   "TT426_4S_ALM_ANALOG_DB_LOW LEVEL VALUE (L)" : Real = PLC TT426_4S_ALM_ANALOG_DB."LOW LEVEL VALUE (L)" AT %DB2080.DBD26, 1 s
   "PIT424PORT_ALM_ANALOG_DB_HIGH LEVEL VALUE (H)" : Real = PLC PIT424PORT_ALM_ANALOG_DB."HIGH LEVEL VALUE (H)" AT %DB2070.DBD30, 1 s
   "TT426_4S_ALM_ANALOG_DB_VERY HIGH LEVEL VALUE (HH)" : Real = PLC TT426_4S_ALM_ANALOG_DB."VERY HIGH LEVEL VALUE (HH)" AT %DB2080.DBD34, 1 s
   "PT415_RIO7_ALM_ANALOG_DB_LOW LEVEL VALUE (L)" : Real = PLC PT415_RIO7_ALM_ANALOG_DB."LOW LEVEL VALUE (L)" AT %DB2225.DBD26, 1 s
   "PT415_RIO6_ALM_ANALOG_DB_VERY HIGH LEVEL VALUE (HH)" : Real = PLC PT415_RIO6_ALM_ANALOG_DB."VERY HIGH LEVEL VALUE (HH)" AT %DB2218.DBD34, 1 s
   "Sequence Times_DB_Pre-Dwell Timer_Days Left" : DInt = PLC "Sequence Times_DB"."Pre-Dwell Timer"."Days Left", 1 s
   "504_Tank Grouping_DB2020_Cycle Period_ET" : Time = PLC "504_Tank Grouping_DB2020"."Cycle Period".ET, 1 s
   "504_Tank Grouping_DB2020_Cycle Length_ET" : Time = PLC "504_Tank Grouping_DB2020"."Cycle Length".ET, 1 s
   "504_Tank Grouping_DB2020_Valve Cycle_Enable" : Bool = PLC "504_Tank Grouping_DB2020"."Valve Cycle".Enable, 1 s
   "504_Tank Grouping_DB2020_Valve Cycle_Period" : Time = PLC "504_Tank Grouping_DB2020"."Valve Cycle".Period, 1 s
   "504_Tank Grouping_DB2020_Valve Cycle_Length" : Time = PLC "504_Tank Grouping_DB2020"."Valve Cycle".Length, 1 s
   "Process Gas Compressor Running/Stopped" : Bool = PLC "Process Gas Compressor Running/Stopped" AT %I139.0, 1 s
   "PT415_FPT_ALM_ANALOG_DB_VERY LOW LEVEL VALUE (LL)" : Real = PLC PT415_FPT_ALM_ANALOG_DB."VERY LOW LEVEL VALUE (LL)" AT %DB2213.DBD22, 1 s
   "PT415_FPT_ALM_ANALOG_DB_LOW LEVEL VALUE (L)" : Real = PLC PT415_FPT_ALM_ANALOG_DB."LOW LEVEL VALUE (L)" AT %DB2213.DBD26, 1 s
   "PT415_FPT_ALM_ANALOG_DB_HIGH LEVEL VALUE (H)" : Real = PLC PT415_FPT_ALM_ANALOG_DB."HIGH LEVEL VALUE (H)" AT %DB2213.DBD30, 1 s
   "PT415_RIO7_ALM_ANALOG_DB_VERY LOW LEVEL VALUE (LL)" : Real = PLC PT415_RIO7_ALM_ANALOG_DB."VERY LOW LEVEL VALUE (LL)" AT %DB2225.DBD22, 1 s
   "PT415_FPT_ALM_ANALOG_DB_VERY HIGH LEVEL VALUE (HH)" : Real = PLC PT415_FPT_ALM_ANALOG_DB."VERY HIGH LEVEL VALUE (HH)" AT %DB2213.DBD34, 1 s
   "PT415_RIO3_ALM_ANALOG_DB_LOW LEVEL VALUE (L)" : Real = PLC PT415_RIO3_ALM_ANALOG_DB."LOW LEVEL VALUE (L)" AT %DB2215.DBD26, 1 s
   "PT415_RIO3_ALM_ANALOG_DB_HIGH LEVEL VALUE (H)" : Real = PLC PT415_RIO3_ALM_ANALOG_DB."HIGH LEVEL VALUE (H)" AT %DB2215.DBD30, 1 s
   "PT415_RIO3_ALM_ANALOG_DB_VERY HIGH LEVEL VALUE (HH)" : Real = PLC PT415_RIO3_ALM_ANALOG_DB."VERY HIGH LEVEL VALUE (HH)" AT %DB2215.DBD34, 1 s
   "PT415_RIO5_ALM_ANALOG_DB_VERY LOW LEVEL VALUE (LL)" : Real = PLC PT415_RIO5_ALM_ANALOG_DB."VERY LOW LEVEL VALUE (LL)" AT %DB2217.DBD22, 1 s
   "PT415_RIO5_ALM_ANALOG_DB_LOW LEVEL VALUE (L)" : Real = PLC PT415_RIO5_ALM_ANALOG_DB."LOW LEVEL VALUE (L)" AT %DB2217.DBD26, 1 s
   "PT415_RIO5_ALM_ANALOG_DB_HIGH LEVEL VALUE (H)" : Real = PLC PT415_RIO5_ALM_ANALOG_DB."HIGH LEVEL VALUE (H)" AT %DB2217.DBD30, 1 s
   "PT415_RIO5_ALM_ANALOG_DB_VERY HIGH LEVEL VALUE (HH)" : Real = PLC PT415_RIO5_ALM_ANALOG_DB."VERY HIGH LEVEL VALUE (HH)" AT %DB2217.DBD34, 1 s
   "PT415_RIO6_ALM_ANALOG_DB_VERY LOW LEVEL VALUE (LL)" : Real = PLC PT415_RIO6_ALM_ANALOG_DB."VERY LOW LEVEL VALUE (LL)" AT %DB2218.DBD22, 1 s
   "PT415_RIO6_ALM_ANALOG_DB_LOW LEVEL VALUE (L)" : Real = PLC PT415_RIO6_ALM_ANALOG_DB."LOW LEVEL VALUE (L)" AT %DB2218.DBD26, 1 s
   "PT415_RIO6_ALM_ANALOG_DB_HIGH LEVEL VALUE (H)" : Real = PLC PT415_RIO6_ALM_ANALOG_DB."HIGH LEVEL VALUE (H)" AT %DB2218.DBD30, 1 s
   "PT415_RIO3_ALM_ANALOG_DB_VERY LOW LEVEL VALUE (LL)" : Real = PLC PT415_RIO3_ALM_ANALOG_DB."VERY LOW LEVEL VALUE (LL)" AT %DB2215.DBD22, 1 s
   "RIO3_SPR_DI_33_4" : Bool = PLC RIO3_SPR_DI_33_4 AT %I33.4, 1 s
   "TT426_1S_ALM_ANALOG_DB_LOW LEVEL VALUE (L)" : Real = PLC TT426_1S_ALM_ANALOG_DB."LOW LEVEL VALUE (L)" AT %DB2076.DBD26, 1 s
   "TT426_1S_ALM_ANALOG_DB_VERY HIGH LEVEL VALUE (HH)" : Real = PLC TT426_1S_ALM_ANALOG_DB."VERY HIGH LEVEL VALUE (HH)" AT %DB2076.DBD34, 1 s
   "RIO6_SPR_DI_66_7" : Bool = PLC RIO6_SPR_DI_66_7 AT %I66.7, 1 s
   "RIO6_SPR_DI_66_5" : Bool = PLC RIO6_SPR_DI_66_5 AT %I66.5, 1 s
   "RIO6_SPR_DI_66_4" : Bool = PLC RIO6_SPR_DI_66_4 AT %I66.4, 1 s
   "RIO6_SPR_DI_66_3" : Bool = PLC RIO6_SPR_DI_66_3 AT %I66.3, 1 s
   "Tank 6S BWT Level High High Switch" : Bool = PLC "Tank 6S BWT Level High High Switch" AT %I66.2, 1 s
   "RIO6 Tanks Pressure Switch Hi Hi" : Bool = PLC "RIO6 Tanks Pressure Switch Hi Hi" AT %I66.1, 1 s
   "Tank 6P BWT Level High High Switch" : Bool = PLC "Tank 6P BWT Level High High Switch" AT %I66.0, 1 s
   "RIO6_SPR_DI_63_7" : Bool = PLC RIO6_SPR_DI_63_7 AT %I63.7, 1 s
   "RIO6_SPR_DI_63_6" : Bool = PLC RIO6_SPR_DI_63_6 AT %I63.6, 1 s
   "Tank 6S Tank Vent Valve 2 Feedback - Closed" : Bool = PLC "Tank 6S Tank Vent Valve 2 Feedback - Closed" AT %I63.5, 1 s
   "Tank 6S Tank Vent Valve 2 Feedback - Opened" : Bool = PLC "Tank 6S Tank Vent Valve 2 Feedback - Opened" AT %I63.4, 1 s
   "Tank 6S Tank Vent Valve 1 Feedback - Closed" : Bool = PLC "Tank 6S Tank Vent Valve 1 Feedback - Closed" AT %I63.3, 1 s
   "Tank 6S Tank Vent Valve 1 Feedback - Opened" : Bool = PLC "Tank 6S Tank Vent Valve 1 Feedback - Opened" AT %I63.2, 1 s
   "Tank 6S GTT Isolation Valve Feedback - Closed" : Bool = PLC "Tank 6S GTT Isolation Valve Feedback - Closed" AT %I63.1, 1 s
   "Tank 6S GTT Isolation Valve Feedback - Opened" : Bool = PLC "Tank 6S GTT Isolation Valve Feedback - Opened" AT %I63.0, 1 s
   "RIO6_SPR_DI_60_7" : Bool = PLC RIO6_SPR_DI_60_7 AT %I60.7, 1 s
   "RIO6_SPR_DI_60_6" : Bool = PLC RIO6_SPR_DI_60_6 AT %I60.6, 1 s
   "Tank 6P Tank Vent Valve 2 Feedback - Closed" : Bool = PLC "Tank 6P Tank Vent Valve 2 Feedback - Closed" AT %I60.5, 1 s
   "Tank 6P Tank Vent Valve 2 Feedback - Opened" : Bool = PLC "Tank 6P Tank Vent Valve 2 Feedback - Opened" AT %I60.4, 1 s
   "Tank 6P Tank Vent Valve 1 Feedback - Closed" : Bool = PLC "Tank 6P Tank Vent Valve 1 Feedback - Closed" AT %I60.3, 1 s
   "Tank 6P Tank Vent Valve 1 Feedback - Opened" : Bool = PLC "Tank 6P Tank Vent Valve 1 Feedback - Opened" AT %I60.2, 1 s
   "RIO6_SPR_DI_66_6" : Bool = PLC RIO6_SPR_DI_66_6 AT %I66.6, 1 s
   "APT GTT Isolation Valve Feedback - Opened" : Bool = PLC "APT GTT Isolation Valve Feedback - Opened" AT %I75.0, 1 s
   "APT GTT Isolation Valve Feedback - Closed" : Bool = PLC "APT GTT Isolation Valve Feedback - Closed" AT %I75.1, 1 s
   "APT Tank Vent Valve 1 Feedback - Opened" : Bool = PLC "APT Tank Vent Valve 1 Feedback - Opened" AT %I75.2, 1 s
   "FIT417_APT_ALM_ANALOG_DB_VERY HIGH LEVEL VALUE (HH)" : Real = PLC FIT417_APT_ALM_ANALOG_DB."VERY HIGH LEVEL VALUE (HH)" AT %DB2099.DBD34, 1 s
   "FIT420_APT_ALM_ANALOG_DB_VERY LOW LEVEL VALUE (LL)" : Real = PLC FIT420_APT_ALM_ANALOG_DB."VERY LOW LEVEL VALUE (LL)" AT %DB2212.DBD22, 1 s
   "FIT420_APT_ALM_ANALOG_DB_LOW LEVEL VALUE (L)" : Real = PLC FIT420_APT_ALM_ANALOG_DB."LOW LEVEL VALUE (L)" AT %DB2212.DBD26, 1 s
   "FIT420_APT_ALM_ANALOG_DB_HIGH LEVEL VALUE (H)" : Real = PLC FIT420_APT_ALM_ANALOG_DB."HIGH LEVEL VALUE (H)" AT %DB2212.DBD30, 1 s
   "FIT420_APT_ALM_ANALOG_DB_VERY HIGH LEVEL VALUE (HH)" : Real = PLC FIT420_APT_ALM_ANALOG_DB."VERY HIGH LEVEL VALUE (HH)" AT %DB2212.DBD34, 1 s
   "TT426_4P_ALM_ANALOG_DB_VERY LOW LEVEL VALUE (LL)" : Real = PLC TT426_4P_ALM_ANALOG_DB."VERY LOW LEVEL VALUE (LL)" AT %DB2079.DBD22, 1 s
   "TT426_4P_ALM_ANALOG_DB_LOW LEVEL VALUE (L)" : Real = PLC TT426_4P_ALM_ANALOG_DB."LOW LEVEL VALUE (L)" AT %DB2079.DBD26, 1 s
   "TT426_4P_ALM_ANALOG_DB_HIGH LEVEL VALUE (H)" : Real = PLC TT426_4P_ALM_ANALOG_DB."HIGH LEVEL VALUE (H)" AT %DB2079.DBD30, 1 s
   "TT426_4P_ALM_ANALOG_DB_VERY HIGH LEVEL VALUE (HH)" : Real = PLC TT426_4P_ALM_ANALOG_DB."VERY HIGH LEVEL VALUE (HH)" AT %DB2079.DBD34, 1 s
   "RIO7_SPR_DI_178_7" : Bool = PLC RIO7_SPR_DI_178_7 AT %I78.7, 1 s
   "Tank 6P GTT Isolation Valve Feedback - Closed" : Bool = PLC "Tank 6P GTT Isolation Valve Feedback - Closed" AT %I60.1, 1 s
   "RIO7_SPR_DI_178_6" : Bool = PLC RIO7_SPR_DI_178_6 AT %I78.6, 1 s
   "RIO7_SPR_DI_178_4" : Bool = PLC RIO7_SPR_DI_178_4 AT %I78.4, 1 s
   "RIO7_SPR_DI_178_3" : Bool = PLC RIO7_SPR_DI_178_3 AT %I78.3, 1 s
   "RIO7_SPR_DI_178_2" : Bool = PLC RIO7_SPR_DI_178_2 AT %I78.2, 1 s
   "RIO7 Tank Pressure Switch Hi Hi" : Bool = PLC "RIO7 Tank Pressure Switch Hi Hi" AT %I78.1, 1 s
   "APT BWT Level High High Switch" : Bool = PLC "APT BWT Level High High Switch" AT %I78.0, 1 s
   "RIO7_SPR_DI_175_7" : Bool = PLC RIO7_SPR_DI_175_7 AT %I75.7, 1 s
   "RIO7_SPR_DI_175_6" : Bool = PLC RIO7_SPR_DI_175_6 AT %I75.6, 1 s
   "APT Tank Vent Valve 2 Feedback - Closed" : Bool = PLC "APT Tank Vent Valve 2 Feedback - Closed" AT %I75.5, 1 s
   "APT Tank Vent Valve 2 Feedback - Opened" : Bool = PLC "APT Tank Vent Valve 2 Feedback - Opened" AT %I75.4, 1 s
   "APT Tank Vent Valve 1 Feedback - Closed" : Bool = PLC "APT Tank Vent Valve 1 Feedback - Closed" AT %I75.3, 1 s
   "RIO7_SPR_DI_178_5" : Bool = PLC RIO7_SPR_DI_178_5 AT %I78.5, 1 s
   "Tank 6P GTT Isolation Valve Feedback - Opened" : Bool = PLC "Tank 6P GTT Isolation Valve Feedback - Opened" AT %I60.0, 1 s
   "RIO5_SPR_DI_57_7" : Bool = PLC RIO5_SPR_DI_57_7 AT %I57.7, 1 s
   "RIO5_SPR_DI_57_6" : Bool = PLC RIO5_SPR_DI_57_6 AT %I57.6, 1 s
   "RIO4_SPR_DI_145_3" : Bool = PLC RIO4_SPR_DI_145_3 AT %I45.3, 1 s
   "Tank 4S BWT Level High High Switch" : Bool = PLC "Tank 4S BWT Level High High Switch" AT %I45.2, 1 s
   "RIO4 Tanks Pressure Switch Hi Hi" : Bool = PLC "RIO4 Tanks Pressure Switch Hi Hi" AT %I45.1, 1 s
   "Tank 4P BWT Level High High Switch" : Bool = PLC "Tank 4P BWT Level High High Switch" AT %I45.0, 1 s
   "RIO4_SPR_DI_142_7" : Bool = PLC RIO4_SPR_DI_142_7 AT %I42.7, 1 s
   "RIO4_SPR_DI_142_6" : Bool = PLC RIO4_SPR_DI_142_6 AT %I42.6, 1 s
   "Tank 4S Tank Vent Valve 2 Feedback - Closed" : Bool = PLC "Tank 4S Tank Vent Valve 2 Feedback - Closed" AT %I42.5, 1 s
   "Tank 4S Tank Vent Valve 2 Feedback - Opened" : Bool = PLC "Tank 4S Tank Vent Valve 2 Feedback - Opened" AT %I42.4, 1 s
   "Tank 4S Tank Vent Valve 1 Feedback - Closed" : Bool = PLC "Tank 4S Tank Vent Valve 1 Feedback - Closed" AT %I42.3, 1 s
   "Tank 4S Tank Vent Valve 1 Feedback - Opened" : Bool = PLC "Tank 4S Tank Vent Valve 1 Feedback - Opened" AT %I42.2, 1 s
   "RIO4_SPR_DI_145_4" : Bool = PLC RIO4_SPR_DI_145_4 AT %I45.4, 1 s
   "Tank 4S GTT Isolation Valve Feedback - Closed" : Bool = PLC "Tank 4S GTT Isolation Valve Feedback - Closed" AT %I42.1, 1 s
   "RIO4_SPR_DI_139_7" : Bool = PLC RIO4_SPR_DI_139_7 AT %I39.7, 1 s
   "RIO4_SPR_DI_139_6" : Bool = PLC RIO4_SPR_DI_139_6 AT %I39.6, 1 s
   "Tank 4P Tank Vent Valve 2 Feedback - Closed" : Bool = PLC "Tank 4P Tank Vent Valve 2 Feedback - Closed" AT %I39.5, 1 s
   "Tank 4P Tank Vent Valve 2 Feedback - Opened" : Bool = PLC "Tank 4P Tank Vent Valve 2 Feedback - Opened" AT %I39.4, 1 s
   "Tank 4P Tank Vent Valve 1 Feedback - Closed" : Bool = PLC "Tank 4P Tank Vent Valve 1 Feedback - Closed" AT %I39.3, 1 s
   "Tank 4P Tank Vent Valve 1 Feedback - Opened" : Bool = PLC "Tank 4P Tank Vent Valve 1 Feedback - Opened" AT %I39.2, 1 s
   "Tank 4P GTT Isolation Valve Feedback - Closed" : Bool = PLC "Tank 4P GTT Isolation Valve Feedback - Closed" AT %I39.1, 1 s
   "Tank 4P GTT Isolation Valve Feedback - Opened" : Bool = PLC "Tank 4P GTT Isolation Valve Feedback - Opened" AT %I39.0, 1 s
   "RIO3_SPR_DI_33_7" : Bool = PLC RIO3_SPR_DI_33_7 AT %I33.7, 1 s
   "RIO3_SPR_DI_33_6" : Bool = PLC RIO3_SPR_DI_33_6 AT %I33.6, 1 s
   "Tank 4S GTT Isolation Valve Feedback - Opened" : Bool = PLC "Tank 4S GTT Isolation Valve Feedback - Opened" AT %I42.0, 1 s
   "FIT417_APT_ALM_ANALOG_DB_HIGH LEVEL VALUE (H)" : Real = PLC FIT417_APT_ALM_ANALOG_DB."HIGH LEVEL VALUE (H)" AT %DB2099.DBD30, 1 s
   "RIO4_SPR_DI_145_5" : Bool = PLC RIO4_SPR_DI_145_5 AT %I45.5, 1 s
   "RIO4_SPR_DI_145_7" : Bool = PLC RIO4_SPR_DI_145_7 AT %I45.7, 1 s
   "RIO5_SPR_DI_57_5" : Bool = PLC RIO5_SPR_DI_57_5 AT %I57.5, 1 s
   "RIO5_SPR_DI_57_4" : Bool = PLC RIO5_SPR_DI_57_4 AT %I57.4, 1 s
   "RIO5_SPR_DI_57_3" : Bool = PLC RIO5_SPR_DI_57_3 AT %I57.3, 1 s
   "Tank 5S BWT Level High High Switch" : Bool = PLC "Tank 5S BWT Level High High Switch" AT %I57.2, 1 s
   "RIO5 Tanks Pressure Switch Hi Hi" : Bool = PLC "RIO5 Tanks Pressure Switch Hi Hi" AT %I57.1, 1 s
   "Tank 5P BWT Level High High Switch" : Bool = PLC "Tank 5P BWT Level High High Switch" AT %I57.0, 1 s
   "RIO5_SPR_DI_54_7" : Bool = PLC RIO5_SPR_DI_54_7 AT %I54.7, 1 s
   "RIO5_SPR_DI_54_6" : Bool = PLC RIO5_SPR_DI_54_6 AT %I54.6, 1 s
   "Tank 5S Tank Vent Valve 2 Feedback - Closed" : Bool = PLC "Tank 5S Tank Vent Valve 2 Feedback - Closed" AT %I54.5, 1 s
   "Tank 5S Tank Vent Valve 2 Feedback - Opened" : Bool = PLC "Tank 5S Tank Vent Valve 2 Feedback - Opened" AT %I54.4, 1 s
   "RIO4_SPR_DI_145_6" : Bool = PLC RIO4_SPR_DI_145_6 AT %I45.6, 1 s
   "Tank 5S Tank Vent Valve 1 Feedback - Closed" : Bool = PLC "Tank 5S Tank Vent Valve 1 Feedback - Closed" AT %I54.3, 1 s
   "Tank 5S GTT Isolation Valve Feedback - Closed" : Bool = PLC "Tank 5S GTT Isolation Valve Feedback - Closed" AT %I54.1, 1 s
   "Tank 5S GTT Isolation Valve Feedback - Opened" : Bool = PLC "Tank 5S GTT Isolation Valve Feedback - Opened" AT %I54.0, 1 s
   "RIO5_SPR_DI_51_7" : Bool = PLC RIO5_SPR_DI_51_7 AT %I51.7, 1 s
   "RIO5_SPR_DI_51_6" : Bool = PLC RIO5_SPR_DI_51_6 AT %I51.6, 1 s
   "Tank 5P Tank Vent Valve 2 Feedback - Closed" : Bool = PLC "Tank 5P Tank Vent Valve 2 Feedback - Closed" AT %I51.5, 1 s
   "Tank 5P Tank Vent Valve 2 Feedback - Opened" : Bool = PLC "Tank 5P Tank Vent Valve 2 Feedback - Opened" AT %I51.4, 1 s
   "Tank 5P Tank Vent Valve 1 Feedback - Closed" : Bool = PLC "Tank 5P Tank Vent Valve 1 Feedback - Closed" AT %I51.3, 1 s
   "Tank 5P Tank Vent Valve 1 Feedback - Opened" : Bool = PLC "Tank 5P Tank Vent Valve 1 Feedback - Opened" AT %I51.2, 1 s
   "Tank 5P GTT Isolation Valve Feedback - Closed" : Bool = PLC "Tank 5P GTT Isolation Valve Feedback - Closed" AT %I51.1, 1 s
   "Tank 5P GTT Isolation Valve Feedback - Opened" : Bool = PLC "Tank 5P GTT Isolation Valve Feedback - Opened" AT %I51.0, 1 s
   "Tank 5S Tank Vent Valve 1 Feedback - Opened" : Bool = PLC "Tank 5S Tank Vent Valve 1 Feedback - Opened" AT %I54.2, 1 s
   "TT426_1S_ALM_ANALOG_DB_HIGH LEVEL VALUE (H)" : Real = PLC TT426_1S_ALM_ANALOG_DB."HIGH LEVEL VALUE (H)" AT %DB2076.DBD30, 1 s
   "FIT417_APT_ALM_ANALOG_DB_LOW LEVEL VALUE (L)" : Real = PLC FIT417_APT_ALM_ANALOG_DB."LOW LEVEL VALUE (L)" AT %DB2099.DBD26, 1 s
   "FIT420_FPT_ALM_ANALOG_DB_VERY HIGH LEVEL VALUE (HH)" : Real = PLC FIT420_FPT_ALM_ANALOG_DB."VERY HIGH LEVEL VALUE (HH)" AT %DB2201.DBD34, 1 s
   "FIT420_1S_ALM_ANALOG_DB_HIGH LEVEL VALUE (H)" : Real = PLC FIT420_1S_ALM_ANALOG_DB."HIGH LEVEL VALUE (H)" AT %DB2203.DBD30, 1 s
   "FIT420_1S_ALM_ANALOG_DB_VERY HIGH LEVEL VALUE (HH)" : Real = PLC FIT420_1S_ALM_ANALOG_DB."VERY HIGH LEVEL VALUE (HH)" AT %DB2203.DBD34, 1 s
   "FIT420_3P_ALM_ANALOG_DB_VERY LOW LEVEL VALUE (LL)" : Real = PLC FIT420_3P_ALM_ANALOG_DB."VERY LOW LEVEL VALUE (LL)" AT %DB2204.DBD22, 1 s
   "FIT420_3P_ALM_ANALOG_DB_LOW LEVEL VALUE (L)" : Real = PLC FIT420_3P_ALM_ANALOG_DB."LOW LEVEL VALUE (L)" AT %DB2204.DBD26, 1 s
   "FIT420_3P_ALM_ANALOG_DB_HIGH LEVEL VALUE (H)" : Real = PLC FIT420_3P_ALM_ANALOG_DB."HIGH LEVEL VALUE (H)" AT %DB2204.DBD30, 1 s
   "FIT420_3P_ALM_ANALOG_DB_VERY HIGH LEVEL VALUE (HH)" : Real = PLC FIT420_3P_ALM_ANALOG_DB."VERY HIGH LEVEL VALUE (HH)" AT %DB2204.DBD34, 1 s
   "FIT418_3P__ALM_ANALOG_DB_VERY LOW LEVEL VALUE (LL)" : Real = PLC "FIT418_3P__ALM_ANALOG_DB"."VERY LOW LEVEL VALUE (LL)" AT %DB2091.DBD22, 1 s
   "FIT418_3P__ALM_ANALOG_DB_LOW LEVEL VALUE (L)" : Real = PLC "FIT418_3P__ALM_ANALOG_DB"."LOW LEVEL VALUE (L)" AT %DB2091.DBD26, 1 s
   "FIT418_3P__ALM_ANALOG_DB_HIGH LEVEL VALUE (H)" : Real = PLC PIT348_ALM_ANALOG_DB73."LOW LEVEL VALUE (L)" AT %DB2091.DBD30, 1 s
   "FIT418_3P__ALM_ANALOG_DB_VERY HIGH LEVEL VALUE (HH)" : Real = PLC "FIT418_3P__ALM_ANALOG_DB"."VERY HIGH LEVEL VALUE (HH)" AT %DB2091.DBD34, 1 s
   "FIT417_3S_ALM_ANALOG_DB_VERY LOW LEVEL VALUE (LL)" : Real = PLC FIT417_3S_ALM_ANALOG_DB."VERY LOW LEVEL VALUE (LL)" AT %DB2092.DBD22, 1 s
   "FIT417_3S_ALM_ANALOG_DB_LOW LEVEL VALUE (L)" : Real = PLC FIT417_3S_ALM_ANALOG_DB."LOW LEVEL VALUE (L)" AT %DB2092.DBD26, 1 s
   "FIT417_3S_ALM_ANALOG_DB_HIGH LEVEL VALUE (H)" : Real = PLC FIT417_3S_ALM_ANALOG_DB."HIGH LEVEL VALUE (H)" AT %DB2092.DBD30, 1 s
   "FIT417_3S_ALM_ANALOG_DB_VERY HIGH LEVEL VALUE (HH)" : Real = PLC FIT417_3S_ALM_ANALOG_DB."VERY HIGH LEVEL VALUE (HH)" AT %DB2092.DBD34, 1 s
   "FIT420_3S_ALM_ANALOG_DB_VERY LOW LEVEL VALUE (LL)" : Real = PLC FIT420_3S_ALM_ANALOG_DB."VERY LOW LEVEL VALUE (LL)" AT %DB2205.DBD22, 1 s
   "FIT420_3S_ALM_ANALOG_DB_LOW LEVEL VALUE (L)" : Real = PLC FIT420_3S_ALM_ANALOG_DB."LOW LEVEL VALUE (L)" AT %DB2205.DBD26, 1 s
   "FIT420_3S_ALM_ANALOG_DB_HIGH LEVEL VALUE (H)" : Real = PLC FIT420_3S_ALM_ANALOG_DB."HIGH LEVEL VALUE (H)" AT %DB2205.DBD30, 1 s
   "FIT420_3S_ALM_ANALOG_DB_VERY HIGH LEVEL VALUE (HH)" : Real = PLC FIT420_3S_ALM_ANALOG_DB."VERY HIGH LEVEL VALUE (HH)" AT %DB2205.DBD34, 1 s
   "FIT418_4P__ALM_ANALOG_DB_VERY LOW LEVEL VALUE (LL)" : Real = PLC "FIT418_4P__ALM_ANALOG_DB"."VERY LOW LEVEL VALUE (LL)" AT %DB2093.DBD22, 1 s
   "FIT418_4P__ALM_ANALOG_DB_LOW LEVEL VALUE (L)" : Real = PLC "FIT418_4P__ALM_ANALOG_DB"."LOW LEVEL VALUE (L)" AT %DB2093.DBD26, 1 s
   "FIT418_4P__ALM_ANALOG_DB_HIGH LEVEL VALUE (H)" : Real = PLC "FIT418_4P__ALM_ANALOG_DB"."HIGH LEVEL VALUE (H)" AT %DB2093.DBD30, 1 s
   "FIT420_1S_ALM_ANALOG_DB_LOW LEVEL VALUE (L)" : Real = PLC FIT420_1S_ALM_ANALOG_DB."LOW LEVEL VALUE (L)" AT %DB2203.DBD26, 1 s
   "FIT420_1S_ALM_ANALOG_DB_VERY LOW LEVEL VALUE (LL)" : Real = PLC FIT420_1S_ALM_ANALOG_DB."VERY LOW LEVEL VALUE (LL)" AT %DB2203.DBD22, 1 s
   "FIT417_1S__ALM_ANALOG_DB_VERY HIGH LEVEL VALUE (HH)" : Real = PLC "FIT417_1S__ALM_ANALOG_DB"."VERY HIGH LEVEL VALUE (HH)" AT %DB2090.DBD34, 1 s
   "FIT417_1S__ALM_ANALOG_DB_HIGH LEVEL VALUE (H)" : Real = PLC "FIT417_1S__ALM_ANALOG_DB"."HIGH LEVEL VALUE (H)" AT %DB2090.DBD30, 1 s
   "PIT424_RIO1_ALM_ANALOG_DB_VERY LOW LEVEL VALUE (LL)" : Real = PLC PIT424_RIO1_ALM_ANALOG_DB."VERY LOW LEVEL VALUE (LL)" AT %DB2219.DBD22, 1 s
   "PIT424_RIO1_ALM_ANALOG_DB_LOW LEVEL VALUE (L)" : Real = PLC PIT424_RIO1_ALM_ANALOG_DB."LOW LEVEL VALUE (L)" AT %DB2219.DBD26, 1 s
   "PIT424_RIO1_ALM_ANALOG_DB_HIGH LEVEL VALUE (H)" : Real = PLC PIT424_RIO1_ALM_ANALOG_DB."HIGH LEVEL VALUE (H)" AT %DB2219.DBD30, 1 s
   "PIT424_RIO1_ALM_ANALOG_DB_VERY HIGH LEVEL VALUE (HH)" : Real = PLC PIT424_RIO1_ALM_ANALOG_DB."VERY HIGH LEVEL VALUE (HH)" AT %DB2219.DBD34, 1 s
   "TT426_1P_ALM_ANALOG_DB_VERY LOW LEVEL VALUE (LL)" : Real = PLC TT426_1P_ALM_ANALOG_DB."VERY LOW LEVEL VALUE (LL)" AT %DB2075.DBD22, 1 s
   "TT426_1P_ALM_ANALOG_DB_LOW LEVEL VALUE (L)" : Real = PLC TT426_1P_ALM_ANALOG_DB."LOW LEVEL VALUE (L)" AT %DB2075.DBD26, 1 s
   "TT426_1P_ALM_ANALOG_DB_HIGH LEVEL VALUE (H)" : Real = PLC TT426_1P_ALM_ANALOG_DB."HIGH LEVEL VALUE (H)" AT %DB2075.DBD30, 1 s
   "TT426_1P_ALM_ANALOG_DB_VERY HIGH LEVEL VALUE (HH)" : Real = PLC TT426_1P_ALM_ANALOG_DB."VERY HIGH LEVEL VALUE (HH)" AT %DB2075.DBD34, 1 s
   "FIT418_FPT__ALM_ANALOG_DB_VERY LOW LEVEL VALUE (LL)" : Real = PLC "FIT418_FPT__ALM_ANALOG_DB"."VERY LOW LEVEL VALUE (LL)" AT %DB2088.DBD22, 1 s
   "FIT418_FPT__ALM_ANALOG_DB_LOW LEVEL VALUE (L)" : Real = PLC "FIT418_FPT__ALM_ANALOG_DB"."LOW LEVEL VALUE (L)" AT %DB2088.DBD26, 1 s
   "FIT418_4P__ALM_ANALOG_DB_VERY HIGH LEVEL VALUE (HH)" : Real = PLC "FIT418_4P__ALM_ANALOG_DB"."VERY HIGH LEVEL VALUE (HH)" AT %DB2093.DBD34, 1 s
   "FIT418_FPT__ALM_ANALOG_DB_HIGH LEVEL VALUE (H)" : Real = PLC "FIT418_FPT__ALM_ANALOG_DB"."HIGH LEVEL VALUE (H)" AT %DB2088.DBD30, 1 s
   "FIT418_1P__ALM_ANALOG_DB_VERY LOW LEVEL VALUE (LL)" : Real = PLC "FIT418_1P__ALM_ANALOG_DB"."VERY LOW LEVEL VALUE (LL)" AT %DB2089.DBD22, 1 s
   "FIT418_1P__ALM_ANALOG_DB_LOW LEVEL VALUE (L)" : Real = PLC "FIT418_1P__ALM_ANALOG_DB"."LOW LEVEL VALUE (L)" AT %DB2089.DBD26, 1 s
   "FIT418_1P__ALM_ANALOG_DB_HIGH LEVEL VALUE (H)" : Real = PLC "FIT418_1P__ALM_ANALOG_DB"."HIGH LEVEL VALUE (H)" AT %DB2089.DBD30, 1 s
   "FIT418_1P__ALM_ANALOG_DB_VERY HIGH LEVEL VALUE (HH)" : Real = PLC "FIT418_1P__ALM_ANALOG_DB"."VERY HIGH LEVEL VALUE (HH)" AT %DB2089.DBD34, 1 s
   "FIT420_1P_ALM_ANALOG_DB_VERY LOW LEVEL VALUE (LL)" : Real = PLC FIT420_1P_ALM_ANALOG_DB."VERY LOW LEVEL VALUE (LL)" AT %DB2202.DBD22, 1 s
   "FIT420_1P_ALM_ANALOG_DB_LOW LEVEL VALUE (L)" : Real = PLC FIT420_1P_ALM_ANALOG_DB."LOW LEVEL VALUE (L)" AT %DB2202.DBD26, 1 s
   "FIT420_1P_ALM_ANALOG_DB_HIGH LEVEL VALUE (H)" : Real = PLC FIT420_1P_ALM_ANALOG_DB."HIGH LEVEL VALUE (H)" AT %DB2202.DBD30, 1 s
   "FIT420_1P_ALM_ANALOG_DB_VERY HIGH LEVEL VALUE (HH)" : Real = PLC FIT420_1P_ALM_ANALOG_DB."VERY HIGH LEVEL VALUE (HH)" AT %DB2202.DBD34, 1 s
   "FIT417_1S__ALM_ANALOG_DB_VERY LOW LEVEL VALUE (LL)" : Real = PLC "FIT417_1S__ALM_ANALOG_DB"."VERY LOW LEVEL VALUE (LL)" AT %DB2090.DBD22, 1 s
   "FIT417_1S__ALM_ANALOG_DB_LOW LEVEL VALUE (L)" : Real = PLC "FIT417_1S__ALM_ANALOG_DB"."LOW LEVEL VALUE (L)" AT %DB2090.DBD26, 1 s
   "FIT418_FPT__ALM_ANALOG_DB_VERY HIGH LEVEL VALUE (HH)" : Real = PLC "FIT418_FPT__ALM_ANALOG_DB"."VERY HIGH LEVEL VALUE (HH)" AT %DB2088.DBD34, 1 s
   "FIT420_4P_ALM_ANALOG_DB_VERY LOW LEVEL VALUE (LL)" : Real = PLC FIT420_4P_ALM_ANALOG_DB."VERY LOW LEVEL VALUE (LL)" AT %DB2206.DBD22, 1 s
   "FIT420_4P_ALM_ANALOG_DB_LOW LEVEL VALUE (L)" : Real = PLC FIT420_4P_ALM_ANALOG_DB."LOW LEVEL VALUE (L)" AT %DB2206.DBD26, 1 s
   "FIT420_4P_ALM_ANALOG_DB_HIGH LEVEL VALUE (H)" : Real = PLC FIT420_4P_ALM_ANALOG_DB."HIGH LEVEL VALUE (H)" AT %DB2206.DBD30, 1 s
   "FIT420_5S_ALM_ANALOG_DB_LOW LEVEL VALUE (L)" : Real = PLC FIT420_5S_ALM_ANALOG_DB."LOW LEVEL VALUE (L)" AT %DB2209.DBD26, 1 s
   "FIT420_5S_ALM_ANALOG_DB_HIGH LEVEL VALUE (H)" : Real = PLC FIT420_5S_ALM_ANALOG_DB."HIGH LEVEL VALUE (H)" AT %DB2209.DBD30, 1 s
   "FIT420_5S_ALM_ANALOG_DB_VERY HIGH LEVEL VALUE (HH)" : Real = PLC FIT420_5S_ALM_ANALOG_DB."VERY HIGH LEVEL VALUE (HH)" AT %DB2209.DBD34, 1 s
   "FIT418_6P__ALM_ANALOG_DB_VERY LOW LEVEL VALUE (LL)" : Real = PLC "FIT418_6P__ALM_ANALOG_DB"."VERY LOW LEVEL VALUE (LL)" AT %DB2097.DBD22, 1 s
   "FIT418_6P__ALM_ANALOG_DB_LOW LEVEL VALUE (L)" : Real = PLC "FIT418_6P__ALM_ANALOG_DB"."LOW LEVEL VALUE (L)" AT %DB2097.DBD26, 1 s
   "FIT418_6P__ALM_ANALOG_DB_HIGH LEVEL VALUE (H)" : Real = PLC "FIT418_6P__ALM_ANALOG_DB"."HIGH LEVEL VALUE (H)" AT %DB2097.DBD30, 1 s
   "FIT418_6P__ALM_ANALOG_DB_VERY HIGH LEVEL VALUE (HH)" : Real = PLC "FIT418_6P__ALM_ANALOG_DB"."VERY HIGH LEVEL VALUE (HH)" AT %DB2097.DBD34, 1 s
   "FIT420_6P_ALM_ANALOG_DB_VERY LOW LEVEL VALUE (LL)" : Real = PLC FIT420_6P_ALM_ANALOG_DB."VERY LOW LEVEL VALUE (LL)" AT %DB2210.DBD22, 1 s
   "FIT420_6P_ALM_ANALOG_DB_LOW LEVEL VALUE (L)" : Real = PLC FIT420_6P_ALM_ANALOG_DB."LOW LEVEL VALUE (L)" AT %DB2210.DBD26, 1 s
   "FIT420_6P_ALM_ANALOG_DB_HIGH LEVEL VALUE (H)" : Real = PLC FIT420_6P_ALM_ANALOG_DB."HIGH LEVEL VALUE (H)" AT %DB2210.DBD30, 1 s
   "FIT420_5S_ALM_ANALOG_DB_VERY LOW LEVEL VALUE (LL)" : Real = PLC FIT420_5S_ALM_ANALOG_DB."VERY LOW LEVEL VALUE (LL)" AT %DB2209.DBD22, 1 s
   "FIT420_6P_ALM_ANALOG_DB_VERY HIGH LEVEL VALUE (HH)" : Real = PLC FIT420_6P_ALM_ANALOG_DB."VERY HIGH LEVEL VALUE (HH)" AT %DB2210.DBD34, 1 s
   "FIT417_6S_ALM_ANALOG_DB_LOW LEVEL VALUE (L)" : Real = PLC FIT417_6S_ALM_ANALOG_DB."LOW LEVEL VALUE (L)" AT %DB2098.DBD26, 1 s
   "FIT417_6S_ALM_ANALOG_DB_HIGH LEVEL VALUE (H)" : Real = PLC FIT417_6S_ALM_ANALOG_DB."HIGH LEVEL VALUE (H)" AT %DB2098.DBD30, 1 s
   "FIT417_6S_ALM_ANALOG_DB_VERY HIGH LEVEL VALUE (HH)" : Real = PLC FIT417_6S_ALM_ANALOG_DB."VERY HIGH LEVEL VALUE (HH)" AT %DB2098.DBD34, 1 s
   "FIT420_6S_ALM_ANALOG_DB_VERY LOW LEVEL VALUE (LL)" : Real = PLC FIT420_6S_ALM_ANALOG_DB."VERY LOW LEVEL VALUE (LL)" AT %DB2211.DBD22, 1 s
   "FIT420_6S_ALM_ANALOG_DB_LOW LEVEL VALUE (L)" : Real = PLC FIT420_6S_ALM_ANALOG_DB."LOW LEVEL VALUE (L)" AT %DB2211.DBD26, 1 s
   "FIT420_6S_ALM_ANALOG_DB_HIGH LEVEL VALUE (H)" : Real = PLC FIT420_6S_ALM_ANALOG_DB."HIGH LEVEL VALUE (H)" AT %DB2211.DBD30, 1 s
   "FIT420_6S_ALM_ANALOG_DB_VERY HIGH LEVEL VALUE (HH)" : Real = PLC FIT420_6S_ALM_ANALOG_DB."VERY HIGH LEVEL VALUE (HH)" AT %DB2211.DBD34, 1 s
   "FIT420_FPT_ALM_ANALOG_DB_VERY LOW LEVEL VALUE (LL)" : Real = PLC FIT420_FPT_ALM_ANALOG_DB."VERY LOW LEVEL VALUE (LL)" AT %DB2201.DBD22, 1 s
   "FIT420_FPT_ALM_ANALOG_DB_LOW LEVEL VALUE (L)" : Real = PLC FIT420_FPT_ALM_ANALOG_DB."LOW LEVEL VALUE (L)" AT %DB2201.DBD26, 1 s
   "FIT420_FPT_ALM_ANALOG_DB_HIGH LEVEL VALUE (H)" : Real = PLC FIT420_FPT_ALM_ANALOG_DB."HIGH LEVEL VALUE (H)" AT %DB2201.DBD30, 1 s
   "FIT417_6S_ALM_ANALOG_DB_VERY LOW LEVEL VALUE (LL)" : Real = PLC FIT417_6S_ALM_ANALOG_DB."VERY LOW LEVEL VALUE (LL)" AT %DB2098.DBD22, 1 s
   "FIT417_APT_ALM_ANALOG_DB_VERY LOW LEVEL VALUE (LL)" : Real = PLC FIT417_APT_ALM_ANALOG_DB."VERY LOW LEVEL VALUE (LL)" AT %DB2099.DBD22, 1 s
   "FIT417_5S_ALM_ANALOG_DB_VERY HIGH LEVEL VALUE (HH)" : Real = PLC FIT417_5S_ALM_ANALOG_DB."VERY HIGH LEVEL VALUE (HH)" AT %DB2096.DBD34, 1 s
   "FIT417_5S_ALM_ANALOG_DB_LOW LEVEL VALUE (L)" : Real = PLC FIT417_5S_ALM_ANALOG_DB."LOW LEVEL VALUE (L)" AT %DB2096.DBD26, 1 s
   "FIT420_4P_ALM_ANALOG_DB_VERY HIGH LEVEL VALUE (HH)" : Real = PLC FIT420_4P_ALM_ANALOG_DB."VERY HIGH LEVEL VALUE (HH)" AT %DB2206.DBD34, 1 s
   "LT422 4P  TANK LEVEL ALARM_VERY LOW LEVEL VALUE (LL)" : Real = PLC "LT422 4P  TANK LEVEL ALARM"."VERY LOW LEVEL VALUE (LL)" AT %DB2233.DBD22, 1 s
   "LT422 4P  TANK LEVEL ALARM_LOW LEVEL VALUE (L)" : Real = PLC "LT422 4P  TANK LEVEL ALARM"."LOW LEVEL VALUE (L)" AT %DB2233.DBD26, 1 s
   "LT422 4P  TANK LEVEL ALARM_HIGH LEVEL VALUE (H)" : Real = PLC "LT422 4P  TANK LEVEL ALARM"."HIGH LEVEL VALUE (H)" AT %DB2233.DBD30, 1 s
   "LT422 4P  TANK LEVEL ALARM_VERY HIGH LEVEL VALUE (HH)" : Real = PLC "LT422 4P  TANK LEVEL ALARM"."VERY HIGH LEVEL VALUE (HH)" AT %DB2233.DBD34, 1 s
   "FIT417_4S_ALM_ANALOG_DB_VERY LOW LEVEL VALUE (LL)" : Real = PLC FIT417_4S_ALM_ANALOG_DB."VERY LOW LEVEL VALUE (LL)" AT %DB2094.DBD22, 1 s
   "FIT417_4S_ALM_ANALOG_DB_LOW LEVEL VALUE (L)" : Real = PLC FIT417_4S_ALM_ANALOG_DB."LOW LEVEL VALUE (L)" AT %DB2094.DBD26, 1 s
   "FIT417_4S_ALM_ANALOG_DB_HIGH LEVEL VALUE (H)" : Real = PLC FIT417_4S_ALM_ANALOG_DB."HIGH LEVEL VALUE (H)" AT %DB2094.DBD30, 1 s
   "FIT417_4S_ALM_ANALOG_DB_VERY HIGH LEVEL VALUE (HH)" : Real = PLC FIT417_4S_ALM_ANALOG_DB."VERY HIGH LEVEL VALUE (HH)" AT %DB2094.DBD34, 1 s
   "FIT420_4S_ALM_ANALOG_DB_VERY LOW LEVEL VALUE (LL)" : Real = PLC FIT420_4S_ALM_ANALOG_DB."VERY LOW LEVEL VALUE (LL)" AT %DB2207.DBD22, 1 s
   "FIT417_5S_ALM_ANALOG_DB_HIGH LEVEL VALUE (H)" : Real = PLC FIT417_5S_ALM_ANALOG_DB."HIGH LEVEL VALUE (H)" AT %DB2096.DBD30, 1 s
   "FIT420_4S_ALM_ANALOG_DB_LOW LEVEL VALUE (L)" : Real = PLC FIT420_4S_ALM_ANALOG_DB."LOW LEVEL VALUE (L)" AT %DB2207.DBD26, 1 s
   "FIT420_4S_ALM_ANALOG_DB_VERY HIGH LEVEL VALUE (HH)" : Real = PLC FIT420_4S_ALM_ANALOG_DB."VERY HIGH LEVEL VALUE (HH)" AT %DB2207.DBD34, 1 s
   "FIT420_5P_ALM_ANALOG_DB_VERY LOW LEVEL VALUE (LL)" : Real = PLC FIT420_5P_ALM_ANALOG_DB."VERY LOW LEVEL VALUE (LL)" AT %DB2208.DBD22, 1 s
   "FIT420_5P_ALM_ANALOG_DB_LOW LEVEL VALUE (L)" : Real = PLC FIT420_5P_ALM_ANALOG_DB."LOW LEVEL VALUE (L)" AT %DB2208.DBD26, 1 s
   "FIT420_5P_ALM_ANALOG_DB_HIGH LEVEL VALUE (H)" : Real = PLC PIT424_RIO1_ALM_ANALOG_DB."LOW LEVEL VALUE (L)" AT %DB2208.DBD30, 1 s
   "FIT420_5P_ALM_ANALOG_DB_VERY HIGH LEVEL VALUE (HH)" : Real = PLC FIT420_5P_ALM_ANALOG_DB."VERY HIGH LEVEL VALUE (HH)" AT %DB2208.DBD34, 1 s
   "FIT418_5P__ALM_ANALOG_DB_VERY LOW LEVEL VALUE (LL)" : Real = PLC "FIT418_5P__ALM_ANALOG_DB"."VERY LOW LEVEL VALUE (LL)" AT %DB2095.DBD22, 1 s
   "FIT418_5P__ALM_ANALOG_DB_LOW LEVEL VALUE (L)" : Real = PLC "FIT418_5P__ALM_ANALOG_DB"."LOW LEVEL VALUE (L)" AT %DB2095.DBD26, 1 s
   "FIT418_5P__ALM_ANALOG_DB_HIGH LEVEL VALUE (H)" : Real = PLC "FIT418_5P__ALM_ANALOG_DB"."HIGH LEVEL VALUE (H)" AT %DB2095.DBD30, 1 s
   "FIT418_5P__ALM_ANALOG_DB_VERY HIGH LEVEL VALUE (HH)" : Real = PLC "FIT418_5P__ALM_ANALOG_DB"."VERY HIGH LEVEL VALUE (HH)" AT %DB2095.DBD34, 1 s
   "FIT417_5S_ALM_ANALOG_DB_VERY LOW LEVEL VALUE (LL)" : Real = PLC FIT417_5S_ALM_ANALOG_DB."VERY LOW LEVEL VALUE (LL)" AT %DB2096.DBD22, 1 s
   "FIT420_4S_ALM_ANALOG_DB_HIGH LEVEL VALUE (H)" : Real = PLC FIT420_4S_ALM_ANALOG_DB."HIGH LEVEL VALUE (H)" AT %DB2207.DBD30, 1 s
   "86_Times_LIT304 Delay" : Time = PLC "86_Times"."LIT304 Delay", 1 s
   "504_Tank Grouping_DB2020_Boost" : Bool = PLC "504_Tank Grouping_DB2020".Boost, 1 s
   "86_Times_P301_START_DLY" : Time = PLC "86_Times".P301_START_DLY, 1 s
   "84_Setpoints_PIT353_InitialFill_Low" : Real = PLC "84_Setpoints".PIT353_InitialFill_Low, 1 s
   "84_Setpoints_PIT353_InitialFill_High" : Real = PLC "84_Setpoints".PIT353_InitialFill_High, 1 s
   "84_Setpoints_PIT353_InitialFill_HighHigh" : Real = PLC "84_Setpoints".PIT353_InitialFill_HighHigh, 1 s
   "84_Setpoints_PIT353_Refill_LowLow" : Real = PLC "84_Setpoints".PIT353_Refill_LowLow, 1 s
   "84_Setpoints_PIT353_Refill_Low" : Real = PLC "84_Setpoints".PIT353_Refill_Low, 1 s
   "84_Setpoints_PIT353_Refill_High" : Real = PLC "84_Setpoints".PIT353_Refill_High, 1 s
   "84_Setpoints_PIT353_Refill_HighHigh" : Real = PLC "84_Setpoints".PIT353_Refill_HighHigh, 1 s
   "82_To_HMI_CRNT_MODE_GCU" : Int = PLC "82_To_HMI".CRNT_MODE_GCU, 1 s
   "80_From_HMI_MAN_DQ_136_0" : Bool = PLC "80_From_HMI".MAN_DQ_136_0, 1 s
   "80_From_HMI_MAN_DQ_136_1" : Bool = PLC "80_From_HMI".MAN_DQ_136_1, 1 s
   "80_From_HMI_MAN_DQ_136_2" : Bool = PLC "80_From_HMI".MAN_DQ_136_2, 1 s
   "80_From_HMI_MAN_DQ_136_3" : Bool = PLC "80_From_HMI".MAN_DQ_136_3, 1 s
   "80_From_HMI_MAN_DQ_136_4" : Bool = PLC "80_From_HMI".MAN_DQ_136_4, 1 s
   "84_Setpoints_PIT353_InitialFill_LowLow" : Real = PLC "84_Setpoints".PIT353_InitialFill_LowLow, 1 s
   "80_From_HMI_MAN_DQ_136_5" : Bool = PLC "80_From_HMI".MAN_DQ_136_5, 1 s
   "80_From_HMI_MAN_DQ_136_7" : Bool = PLC "80_From_HMI".MAN_DQ_136_7, 1 s
   "80_From_HMI_MAN_DQ_137_0" : Bool = PLC "80_From_HMI".MAN_DQ_137_0, 1 s
   "80_From_HMI_MAN_DQ_137_1" : Bool = PLC "80_From_HMI".MAN_DQ_137_1, 1 s
   "80_From_HMI_MAN_DQ_137_2" : Bool = PLC "80_From_HMI".MAN_DQ_137_2, 1 s
   "80_From_HMI_MAN_DQ_137_3" : Bool = PLC "80_From_HMI".MAN_DQ_137_3, 1 s
   "80_From_HMI_MAN_DQ_137_4" : Bool = PLC "80_From_HMI".MAN_DQ_137_4, 1 s
   "80_From_HMI_MAN_DQ_137_5" : Bool = PLC "80_From_HMI".MAN_DQ_137_5, 1 s
   "80_From_HMI_MAN_DQ_137_6" : Bool = PLC "80_From_HMI".MAN_DQ_137_6, 1 s
   "80_From_HMI_MAN_DQ_137_7" : Bool = PLC "80_From_HMI".MAN_DQ_137_7, 1 s
   "80_From_HMI_MAN_DQ_138_0" : Bool = PLC "80_From_HMI".MAN_DQ_138_0, 1 s
   "80_From_HMI_MAN_DQ_138_1" : Bool = PLC "80_From_HMI".MAN_DQ_138_1, 1 s
   "80_From_HMI_MAN_DQ_138_2" : Bool = PLC "80_From_HMI".MAN_DQ_138_2, 1 s
   "80_From_HMI_MAN_DQ_138_3" : Bool = PLC "80_From_HMI".MAN_DQ_138_3, 1 s
   "80_From_HMI_MAN_DQ_136_6" : Bool = PLC "80_From_HMI".MAN_DQ_136_6, 1 s
   "80_From_HMI_MAN_DQ_138_4" : Bool = PLC "80_From_HMI".MAN_DQ_138_4, 1 s
   "84_Setpoints_PIT358_Refill_HighHigh" : Real = PLC "84_Setpoints".PIT358_Refill_HighHigh, 1 s
   "84_Setpoints_PIT358_Refill_Low" : Real = PLC "84_Setpoints".PIT358_Refill_Low, 1 s
   "84_Setpoints_PIT416_High" : Real = PLC "84_Setpoints".PIT416_High, 1 s
   "19_AUTO_CMNDS_Data_PIT358_CMND_LowLow" : Real = PLC "19_AUTO_CMNDS_Data".PIT358_CMND_LowLow, 1 s
   "19_AUTO_CMNDS_Data_PIT358_CMND_Low" : Real = PLC "19_AUTO_CMNDS_Data".PIT358_CMND_Low, 1 s
   "19_AUTO_CMNDS_Data_PIT358_CMND_High" : Real = PLC "19_AUTO_CMNDS_Data".PIT358_CMND_High, 1 s
   "19_AUTO_CMNDS_Data_PIT358_CMND_HighHigh" : Real = PLC "19_AUTO_CMNDS_Data".PIT358_CMND_HighHigh, 1 s
   "84_Setpoints_PIT348_LowLow" : Real = PLC "84_Setpoints".PIT348_LowLow, 1 s
   "84_Setpoints_PIT348_Low" : Real = PLC "84_Setpoints".PIT348_Low, 1 s
   "84_Setpoints_PIT348_High" : Real = PLC "84_Setpoints".PIT348_High, 1 s
   "84_Setpoints_PIT348_HighHigh" : Real = PLC "84_Setpoints".PIT348_HighHigh, 1 s
   "84_Setpoints_E400_PT002_High" : Real = PLC "84_Setpoints".E400_PT002_High, 1 s
   "84_Setpoints_E400_TT002_High" : Real = PLC "84_Setpoints".E400_TT002_High, 1 s
   "19_AUTO_CMNDS_Data_PIT353_CMND_LowLow" : Real = PLC "19_AUTO_CMNDS_Data".PIT353_CMND_LowLow, 1 s
   "19_AUTO_CMNDS_Data_PIT353_CMND_Low" : Real = PLC "19_AUTO_CMNDS_Data".PIT353_CMND_Low, 1 s
   "84_Setpoints_PIT358_Refill_High" : Real = PLC "84_Setpoints".PIT358_Refill_High, 1 s
   "19_AUTO_CMNDS_Data_PIT353_CMND_High" : Real = PLC "19_AUTO_CMNDS_Data".PIT353_CMND_High, 1 s
   "84_Setpoints_LIT304_InitialFill_LowLow" : Real = PLC "84_Setpoints".LIT304_InitialFill_LowLow, 1 s
   "84_Setpoints_LIT304_InitialFill_Target" : Real = PLC "84_Setpoints".LIT304_InitialFill_Target, 1 s
   "84_Setpoints_LIT304_InitialFill_HighHigh" : Real = PLC "84_Setpoints".LIT304_InitialFill_HighHigh, 1 s
   "84_Setpoints_LIT304_Refill_LowLow" : Real = PLC "84_Setpoints".LIT304_Refill_LowLow, 1 s
   "84_Setpoints_LIT304_Refill_Low" : Real = PLC "84_Setpoints".LIT304_Refill_Low, 1 s
   "84_Setpoints_LIT304_Refill_Target" : Real = PLC "84_Setpoints".LIT304_Refill_Target, 1 s
